// TIA Portal project "HydroPlantProject_V15.1" (V15.1) (continued)

   IF "StationIntHoa" = 1 OR ("StationIntHoa" = 2 AND "StationIntl_Ctrl") THEN
       "StationInterlock_Out" := 1;
   END_IF;

   IF "BaffleHOA" = 0 OR ("BaffleHOA" = 2 AND NOT "Baffle_Ctrl") THEN
       "Baffle_En" := 0;
   END_IF;

   IF "BaffleHOA" = 1 OR ("BaffleHOA" = 2 AND "Baffle_Ctrl") THEN
       "Baffle_En" := 1;
   END_IF;





   //Analog Outputs
   "SCP"(Input_Min:=0,
         Input_Signal:="OilPumpVFDpct",
         Input_Max:=100,
         Output_Min:=0,
         Output_Max:=27648,
         SV=>"OilPumpVFDsp_Out");

   "SCP"(Input_Min := 0,
         Input_Signal := "BafflePct",
         Input_Max := 100,
         Output_Min := 0,
         Output_Max := 27648,
         SV => "Baffle_Out");


   //Analog Inputs
   "SCP"(Input_Min:=0,
         Input_Signal:="OilTemp_In",
         Input_Max:=27648,
         Output_Min:=0,
         Output_Max:=500,
         SV=>"OilTemp");

   "SCP"(Input_Min := 0,
         Input_Signal := "OilFlow_In",
         Input_Max := 27648,
         Output_Min := 0,
         Output_Max := 30,
         SV => "OilFlow");

   "SCP"(Input_Min := 0,
         Input_Signal := "RPM_In",
   Input_Max := 27648,
   Output_Min := 0,
   Output_Max := 200,
   SV => "RPM");

   "SCP"(Input_Min := 0,
         Input_Signal := "Current_In",
         Input_Max := 27648,
         Output_Min := 0,
         Output_Max := 700,
         SV => "Current");


   //Full Auto Bit
   IF "BaffleHOA" = 2 AND "AlarmHornHoa" = 0 AND "VFDHOA" = 0 AND "StationIntHoa" = 0 AND "BrakeHoa" = 0 THEN
       "FullAutoBit" := 1;
   ELSE
       "FullAutoBit" := 0;
   END_IF;
END_FUNCTION_BLOCK

FUNCTION_BLOCK "IO_STL"   // FB5, STL
{ S7_Optimized_Access := 'TRUE' }
VERSION : 0.1
BEGIN

REGION Network 1
   //Digital Outputs
         A     "OilLowFlowAlarm";
         JC    ResetOilPumpVFD;
         CLR;
         A     "EStopAlarm";
         JC    ResetOilPumpVFD;
         L     "VFDHOA";
         L     0;
         ==I;
         JC    ResetOilPumpVFD;
         CLR;
         L     "VFDHOA";
         L     1;
         ==I;
         JC    SetOilPumpVFD;
         CLR;
         L     "VFDHOA";
         L     2;
         ==I;
         JC    AutoOilPumpVFD;

   AutoOilPumpVFD:A     "OilPumpVFD_Ctrl";
         JC    SetOilPumpVFD;
         JU    ResetOilPumpVFD;

   SetOilPumpVFD:AN    "OilLowFlowAlarm";
         AN    "EStop";
         S     "OilPumpVFDen_Out";
         JU    Brake;

   ResetOilPumpVFD:R     "OilPumpVFDen_Out";
         JU    Brake;

   Brake:L     "BrakeHoa";
         L     0;
         ==I;
         JC    ResetBrake;
         CLR;
         L     "BrakeHoa";
         L     1;
         ==I;
         JC    SetBrake;
         CLR;
         L     "BrakeHoa";
         L     2;
         ==I;
         JC    AutoBrake;

   AutoBrake:A     "Brake_Ctrl";
         JC    SetBrake;
         JU    ResetBrake;

   SetBrake:S     "Brake_Out";
         JU    AlarmHorn;

   ResetBrake:R     "Brake_Out";
         JU    AlarmHorn;

   AlarmHorn:L     "AlarmHornHoa";
         L     0;
         ==I;
         JC    ResetAlarmHorn;
         CLR;
         L     "AlarmHornHoa";
         L     1;
         ==I;
         JC    SetAlarmHorn;
         CLR;
         L     "AlarmHornHoa";
         L     2;
         ==I;
         JC    AutoAlarmHorn;

   AutoAlarmHorn:A     "AlarmHorn_Ctrl";
         JC    SetAlarmHorn;
         JU    ResetAlarmHorn;

   SetAlarmHorn:S     "AlarmHorn_Out";
         JU    StationInterlock;

   ResetAlarmHorn:R     "AlarmHorn_Out";
         JU    StationInterlock;

   StationInterlock:A     "EStopAlarm";
         JC    ResetStationInterlock;
         L     "StationIntHoa";
         L     0;
         ==I;
         JC    ResetStationInterlock;
         CLR;
         L     "StationIntHoa";
         L     1;
         ==I;
         JC    SetStationInterlock;
         CLR;
         L     "StationIntHoa";
         L     2;
         ==I;
         JC    AutoStationInterlock;

   AutoStationInterlock:A     "StationIntl_Ctrl";
         JC    SetStationInterlock;
         JU    ResetStationInterlock;

   SetStationInterlock:AN    "EStopAlarm";
         S     "StationInterlock_Out";
         JU    Baffle;

   ResetStationInterlock:R     "StationInterlock_Out";
         JU    Baffle;

   Baffle:L     "BaffleHOA";
         L     0;
         ==I;
         JC    ResetBaffle;
         CLR;
         L     "BaffleHOA";
         L     1;
         ==I;
         JC    SetBaffle;
         CLR;
         L     "BaffleHOA";
         L     2;
         ==I;
         JC    AutoBaffle;

   AutoBaffle:A     "Baffle_Ctrl";
         JC    SetBaffle;
         JU    ResetBaffle;

   SetBaffle:S     "Baffle_En";
         JU    AnalogOutputs;

   ResetBaffle:R     "Baffle_En";
         JU    AnalogOutputs;



   //Analog Outputs
   AnalogOutputs:CALL  "SCP"
         ( Input_Min    := 0,
           Input_Signal := "OilPumpVFDpct",
           Input_Max    := 100,
           Output_Min   := 0,
           Output_Max   := 27648,
           SV           := "OilPumpVFDsp_Out"
         );
         JU    AnalogInputs;

         CALL  "SCP"
         ( Input_Min    := 0,
           Input_Signal := "BafflePct",
           Input_Max    := 100,
           Output_Min   := 0,
           Output_Max   := 27648,
           SV           := "Baffle_Out"
         );


   //Analog Inputs
   AnalogInputs:CALL  "SCP"
         ( Input_Min    := 0,
           Input_Signal := "OilTemp_In",
           Input_Max    := 27648,
           Output_Min   := 0,
           Output_Max   := 500,
           SV           := "OilTemp"
         );

         CALL  "SCP"
         ( Input_Min    := 0,
           Input_Signal := "OilFlow_In",
           Input_Max    := 27648,
           Output_Min   := 0,
           Output_Max   := 30,
           SV           := "OilFlow"
         );

         CALL  "SCP"
         ( Input_Min    := 0,
           Input_Signal := "RPM_In",
           Input_Max    := 27648,
           Output_Min   := 0,
           Output_Max   := 200,
           SV           := "RPM"
         );

         CALL  "SCP"
         ( Input_Min    := 0,
           Input_Signal := "Current_In",
           Input_Max    := 27648,
           Output_Min   := 0,
           Output_Max   := 700,
           SV           := "Current"
         );

   //Full Auto Bit
         CLR;
         L     "BaffleHOA";
         L     2;
         ==I;
         NOT;
         JC    ResetFullAuto;
         CLR;
         L     "VFDHOA";
         L     2;
         ==I;
         NOT;
         JC    ResetFullAuto;
         CLR;
         L     "AlarmHornHoa";
         L     2;
         ==I;
         NOT;
         JC    ResetFullAuto;
         CLR;
         L     "BrakeHoa";
         L     2;
         ==I;
         NOT;
         JC    ResetFullAuto;
         CLR;
         L     "StationIntHoa";
         L     2;
         ==I;
         NOT;
         JC    ResetFullAuto;
         CLR;
         SET;
         S     "FullAutoBit";
         JU    EndOfLine;

   ResetFullAuto:SET;
         NOT;
         R     "FullAutoBit";
         JU    EndOfLine;

   EndOfLine:BE;
END_REGION
END_FUNCTION_BLOCK

FUNCTION_BLOCK "ALARMS_LAD"   // FB6, LAD
{ S7_Optimized_Access := 'TRUE' }
VERSION : 0.1
   VAR
      OS1 : Bool;
      OS2 : Bool;
      OS3 : Bool;
      OS4 : Bool;
      OS5 : Bool;
      OS6 : Bool;
      OS7 : Bool;
      OS8 : Bool;
   END_VAR
   VAR_TEMP
      tv : Time;
      Tsp : Int;
      OLFAT : Bool;
      OLFD : Int;
      tv1 : Time;
      OCD : Int;
      tv2 : Time;
      OCAT : Bool;
      HOTD : Int;
      tv3 : Time;
      HOTAT : Bool;
      OSD : Int;
      tv4 : Time;
      OSAT : Bool;
      OHFD : Int;
      tv5 : Time;
      OHFAT : Bool;
      BFD : Int;
      tv6 : Time;
      BFAT : Bool;
      ESAT : Bool;
      AlarmHornTrigger : Bool;
   END_VAR
   VAR_TEMP   // added for the SCL form of the ladder/FBD networks
      _w1 : Bool;
      _w2 : Bool;
   END_VAR
BEGIN

REGION Network 1
   // Oil Low Flow Alarm
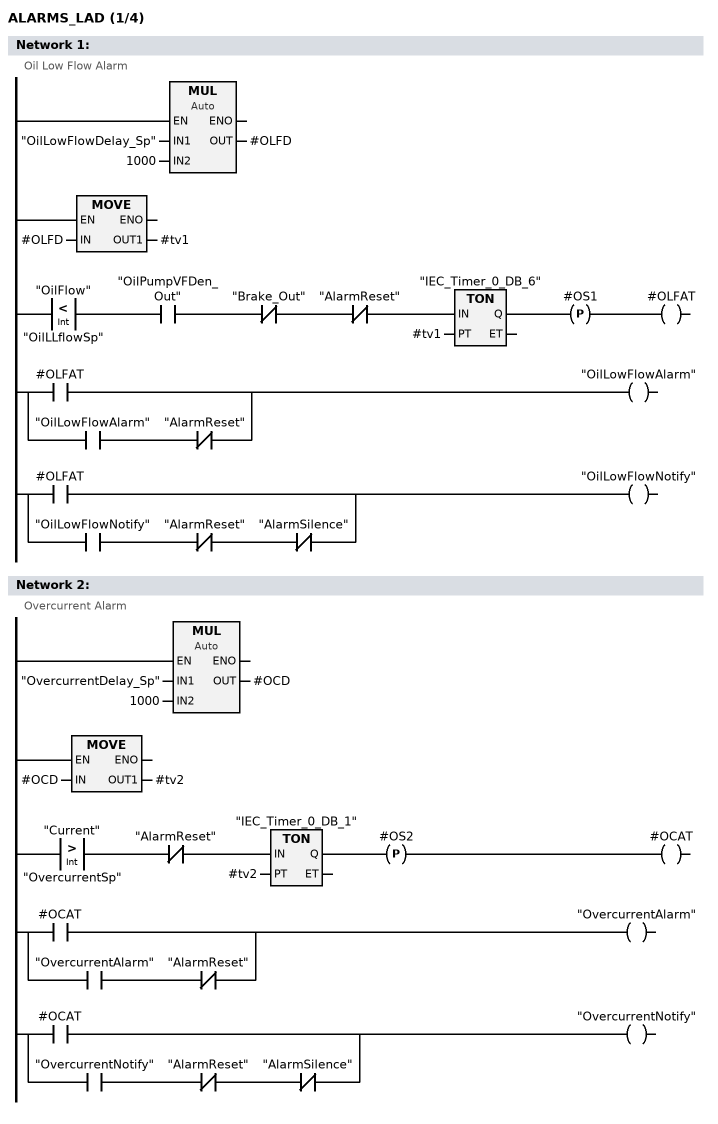
   #OLFD := "OilLowFlowDelay_Sp" * 1000;
   #tv1 := #OLFD;
   "IEC_Timer_0_DB_6".TON(IN := ("OilFlow" < "OilLLflowSp") AND "OilPumpVFDen_Out" AND NOT "Brake_Out" AND NOT "AlarmReset",
                          PT := #tv1);
   #_w1 := "IEC_Timer_0_DB_6".Q AND NOT #OS1;   // rising edge
   #OS1 := "IEC_Timer_0_DB_6".Q;
   #OLFAT := #_w1;
   "OilLowFlowAlarm" := #OLFAT OR ("OilLowFlowAlarm" AND NOT "AlarmReset");
   "OilLowFlowNotify" := #OLFAT OR ("OilLowFlowNotify" AND NOT "AlarmReset" AND NOT "AlarmSilence");
END_REGION

REGION Network 2
   // Overcurrent Alarm
   #OCD := "OvercurrentDelay_Sp" * 1000;
   #tv2 := #OCD;
   "IEC_Timer_0_DB_1".TON(IN := ("Current" > "OvercurrentSp") AND NOT "AlarmReset", PT := #tv2);
   #_w1 := "IEC_Timer_0_DB_1".Q AND NOT #OS2;   // rising edge
   #OS2 := "IEC_Timer_0_DB_1".Q;
   #OCAT := #_w1;
   "OvercurrentAlarm" := #OCAT OR ("OvercurrentAlarm" AND NOT "AlarmReset");
   "OvercurrentNotify" := #OCAT OR ("OvercurrentNotify" AND NOT "AlarmReset" AND NOT "AlarmSilence");
END_REGION

REGION Network 3
   // High Oil Temp Alarm
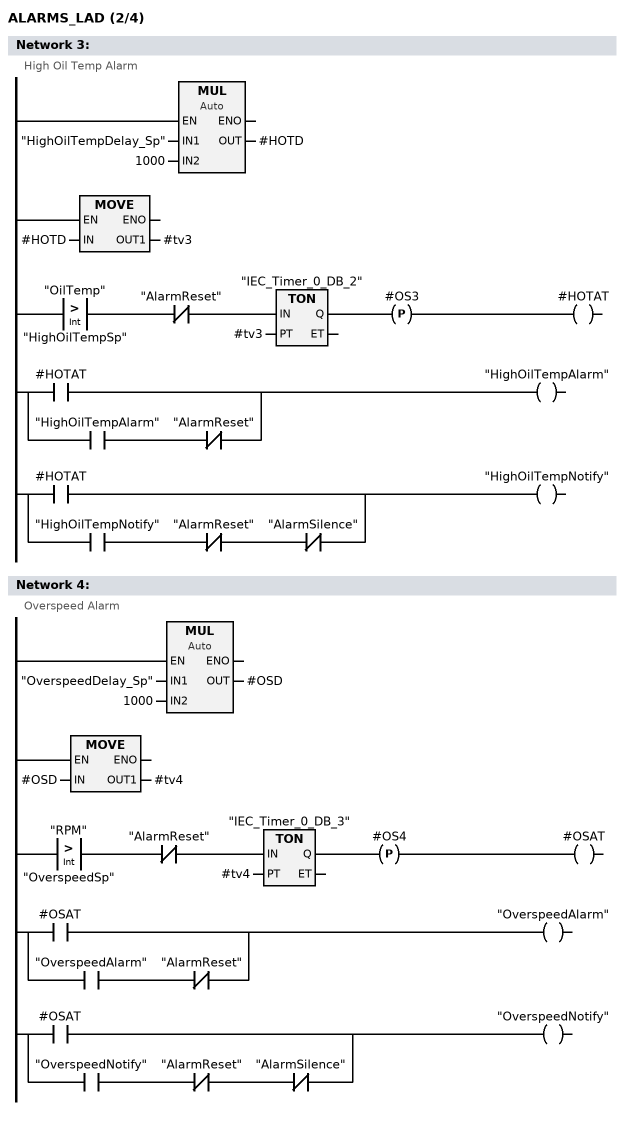
   #HOTD := "HighOilTempDelay_Sp" * 1000;
   #tv3 := #HOTD;
   "IEC_Timer_0_DB_2".TON(IN := ("OilTemp" > "HighOilTempSp") AND NOT "AlarmReset", PT := #tv3);
   #_w1 := "IEC_Timer_0_DB_2".Q AND NOT #OS3;   // rising edge
   #OS3 := "IEC_Timer_0_DB_2".Q;
   #HOTAT := #_w1;
   "HighOilTempAlarm" := #HOTAT OR ("HighOilTempAlarm" AND NOT "AlarmReset");
   "HighOilTempNotify" := #HOTAT OR ("HighOilTempNotify" AND NOT "AlarmReset" AND NOT "AlarmSilence");
END_REGION

REGION Network 4
   // Overspeed Alarm
   #OSD := "OverspeedDelay_Sp" * 1000;
   #tv4 := #OSD;
   "IEC_Timer_0_DB_3".TON(IN := ("RPM" > "OverspeedSp") AND NOT "AlarmReset", PT := #tv4);
   #_w1 := "IEC_Timer_0_DB_3".Q AND NOT #OS4;   // rising edge
   #OS4 := "IEC_Timer_0_DB_3".Q;
   #OSAT := #_w1;
   "OverspeedAlarm" := #OSAT OR ("OverspeedAlarm" AND NOT "AlarmReset");
   "OverspeedNotify" := #OSAT OR ("OverspeedNotify" AND NOT "AlarmReset" AND NOT "AlarmSilence");
END_REGION

REGION Network 5
   // Oil High Flow Alarm
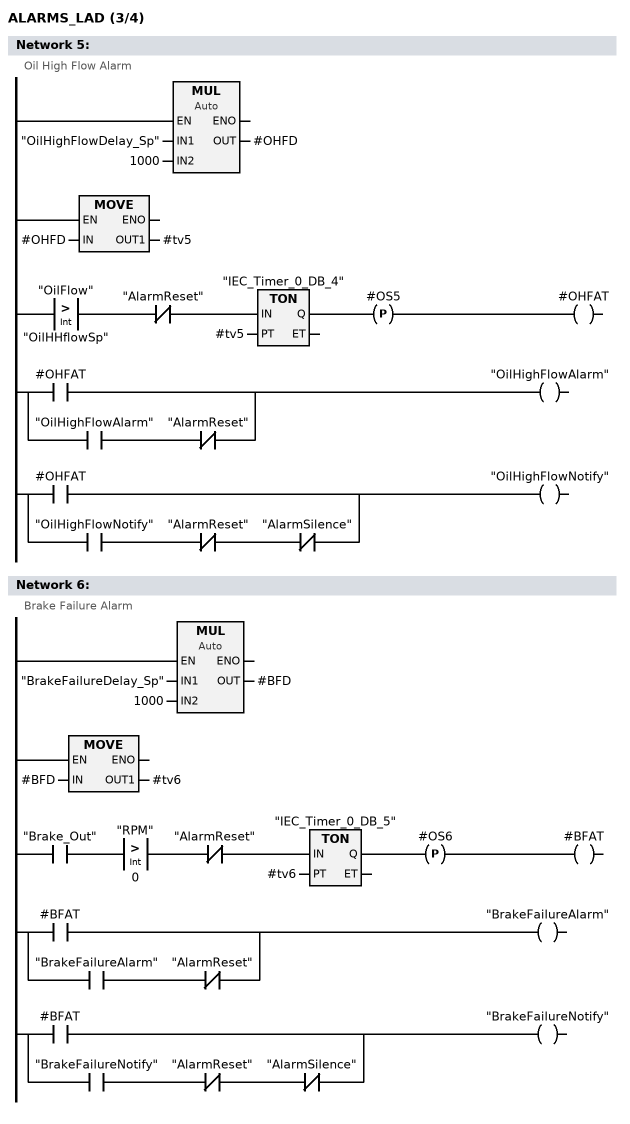
   #OHFD := "OilHighFlowDelay_Sp" * 1000;
   #tv5 := #OHFD;
   "IEC_Timer_0_DB_4".TON(IN := ("OilFlow" > "OilHHflowSp") AND NOT "AlarmReset", PT := #tv5);
   #_w1 := "IEC_Timer_0_DB_4".Q AND NOT #OS5;   // rising edge
   #OS5 := "IEC_Timer_0_DB_4".Q;
   #OHFAT := #_w1;
   "OilHighFlowAlarm" := #OHFAT OR ("OilHighFlowAlarm" AND NOT "AlarmReset");
   "OilHighFlowNotify" := #OHFAT OR ("OilHighFlowNotify" AND NOT "AlarmReset" AND NOT "AlarmSilence");
END_REGION

REGION Network 6
   // Brake Failure Alarm
   #BFD := "BrakeFailureDelay_Sp" * 1000;
   #tv6 := #BFD;
   "IEC_Timer_0_DB_5".TON(IN := "Brake_Out" AND ("RPM" > 0) AND NOT "AlarmReset", PT := #tv6);
   #_w1 := "IEC_Timer_0_DB_5".Q AND NOT #OS6;   // rising edge
   #OS6 := "IEC_Timer_0_DB_5".Q;
   #BFAT := #_w1;
   "BrakeFailureAlarm" := #BFAT OR ("BrakeFailureAlarm" AND NOT "AlarmReset");
   "BrakeFailureNotify" := #BFAT OR ("BrakeFailureNotify" AND NOT "AlarmReset" AND NOT "AlarmSilence");
END_REGION

REGION Network 7
   // EStop Alarm
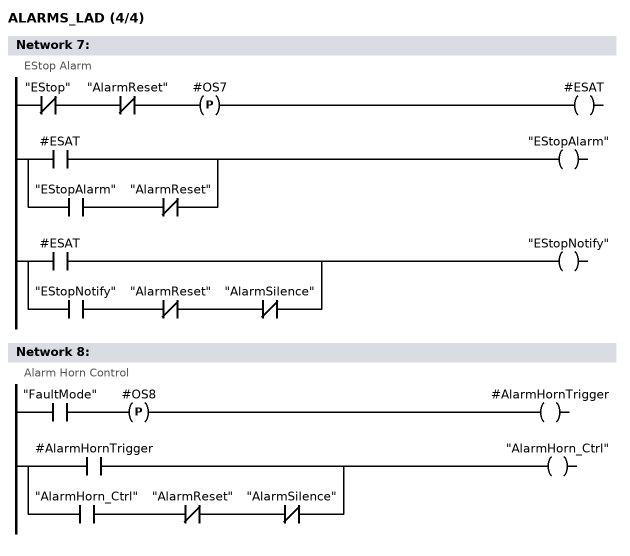
   RUNG wire#powerrail
      I_Contact( "EStop" )
      I_Contact( "AlarmReset" )
      P_Trig( #OS7 )
      Coil( #ESAT )
   END_RUNG
   RUNG wire#powerrail
      Contact( #ESAT )
      wire#w1
      Coil( "EStopAlarm" )
   END_RUNG
   RUNG wire#powerrail
      Contact( "EStopAlarm" )
      I_Contact( "AlarmReset" )
   END_RUNG wire#w1
   RUNG wire#powerrail
      Contact( #ESAT )
      wire#w2
      Coil( "EStopNotify" )
   END_RUNG
   RUNG wire#powerrail
      Contact( "EStopNotify" )
      I_Contact( "AlarmReset" )
      I_Contact( "AlarmSilence" )
   END_RUNG wire#w2
   // the same network as SCL:
   #_w1 := NOT "EStop" AND NOT "AlarmReset";
   #_w2 := #_w1 AND NOT #OS7;   // rising edge
   #OS7 := #_w1;
   #ESAT := #_w2;
   "EStopAlarm" := #ESAT OR ("EStopAlarm" AND NOT "AlarmReset");
   "EStopNotify" := #ESAT OR ("EStopNotify" AND NOT "AlarmReset" AND NOT "AlarmSilence");
END_REGION

REGION Network 8
   // Alarm Horn Control
   RUNG wire#powerrail
      Contact( "FaultMode" )
      P_Trig( #OS8 )
      Coil( #AlarmHornTrigger )
   END_RUNG
   RUNG wire#powerrail
      Contact( #AlarmHornTrigger )
      wire#w1
      Coil( "AlarmHorn_Ctrl" )
   END_RUNG
   RUNG wire#powerrail
      Contact( "AlarmHorn_Ctrl" )
      I_Contact( "AlarmReset" )
      I_Contact( "AlarmSilence" )
   END_RUNG wire#w1
   // the same network as SCL:
   #_w1 := "FaultMode" AND NOT #OS8;   // rising edge
   #OS8 := "FaultMode";
   #AlarmHornTrigger := #_w1;
   "AlarmHorn_Ctrl" := #AlarmHornTrigger OR ("AlarmHorn_Ctrl" AND NOT "AlarmReset" AND NOT "AlarmSilence");
END_REGION
END_FUNCTION_BLOCK

FUNCTION_BLOCK "HOA_FBD"   // FB7, FBD
{ S7_Optimized_Access := 'TRUE' }
VERSION : 0.1
   VAR
      OS1 : Bool;
      OS3 : Bool;
      OS2 : Bool;
      OS4 : Bool;
      OS5 : Bool;
      OS6 : Bool;
      OS7 : Bool;
      OS8 : Bool;
      OS9 : Bool;
      OS10 : Bool;
      OS11 : Bool;
      OS12 : Bool;
   END_VAR
   VAR_TEMP   // added for the SCL form of the ladder/FBD networks
      _w1 : Bool;
      _w2 : Bool;
      _w3 : Bool;
   END_VAR
BEGIN

REGION Network 1
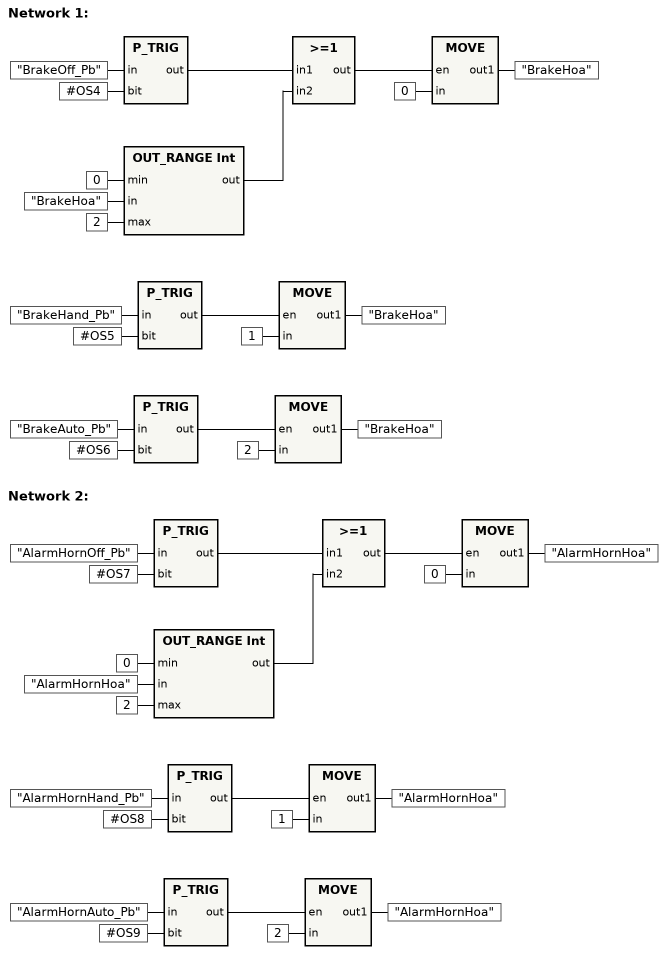
   #_w1 := "BrakeOff_Pb" AND NOT #OS4;   // rising edge
   #OS4 := "BrakeOff_Pb";
   IF #_w1 OR ("BrakeHoa" < 0) OR ("BrakeHoa" > 2) THEN "BrakeHoa" := 0; END_IF;
   #_w2 := "BrakeHand_Pb" AND NOT #OS5;   // rising edge
   #OS5 := "BrakeHand_Pb";
   IF #_w2 THEN "BrakeHoa" := 1; END_IF;
   #_w3 := "BrakeAuto_Pb" AND NOT #OS6;   // rising edge
   #OS6 := "BrakeAuto_Pb";
   IF #_w3 THEN "BrakeHoa" := 2; END_IF;
END_REGION

REGION Network 2
   #_w1 := "AlarmHornOff_Pb" AND NOT #OS7;   // rising edge
   #OS7 := "AlarmHornOff_Pb";
   IF #_w1 OR ("AlarmHornHoa" < 0) OR ("AlarmHornHoa" > 2) THEN "AlarmHornHoa" := 0; END_IF;
   #_w2 := "AlarmHornHand_Pb" AND NOT #OS8;   // rising edge
   #OS8 := "AlarmHornHand_Pb";
   IF #_w2 THEN "AlarmHornHoa" := 1; END_IF;
   #_w3 := "AlarmHornAuto_Pb" AND NOT #OS9;   // rising edge
   #OS9 := "AlarmHornAuto_Pb";
   IF #_w3 THEN "AlarmHornHoa" := 2; END_IF;
END_REGION

REGION Network 3
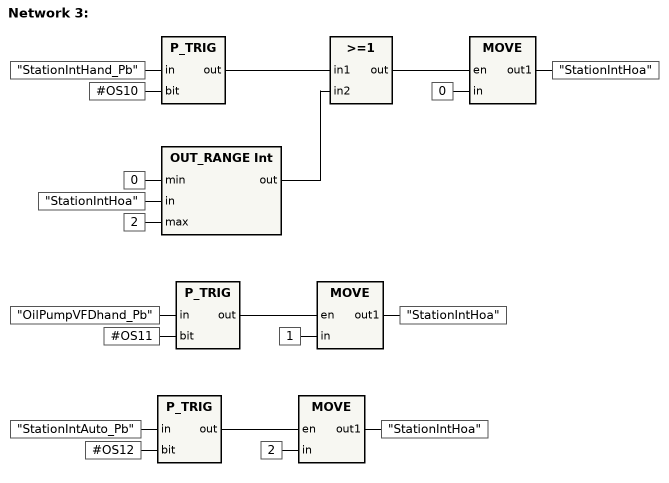
   #_w1 := "StationIntHand_Pb" AND NOT #OS10;   // rising edge
   #OS10 := "StationIntHand_Pb";
   IF #_w1 OR ("StationIntHoa" < 0) OR ("StationIntHoa" > 2) THEN "StationIntHoa" := 0; END_IF;
   #_w2 := "OilPumpVFDhand_Pb" AND NOT #OS11;   // rising edge
   #OS11 := "OilPumpVFDhand_Pb";
   IF #_w2 THEN "StationIntHoa" := 1; END_IF;
   #_w3 := "StationIntAuto_Pb" AND NOT #OS12;   // rising edge
   #OS12 := "StationIntAuto_Pb";
   IF #_w3 THEN "StationIntHoa" := 2; END_IF;
END_REGION
END_FUNCTION_BLOCK

FUNCTION_BLOCK "HOA_LAD"   // FB8, LAD
{ S7_Optimized_Access := 'TRUE' }
VERSION : 0.1
   VAR
      OS1 : Bool;
      OS2 : Bool;
      OS3 : Bool;
      OS4 : Bool;
      OS5 : Bool;
      OS6 : Bool;
      OS7 : Bool;
      OS8 : Bool;
      OS9 : Bool;
      OS10 : Bool;
      OS11 : Bool;
      OS12 : Bool;
   END_VAR
   VAR_TEMP   // added for the SCL form of the ladder/FBD networks
      _w1 : Bool;
      _w2 : Bool;
      _w3 : Bool;
   END_VAR
BEGIN

REGION Network 1
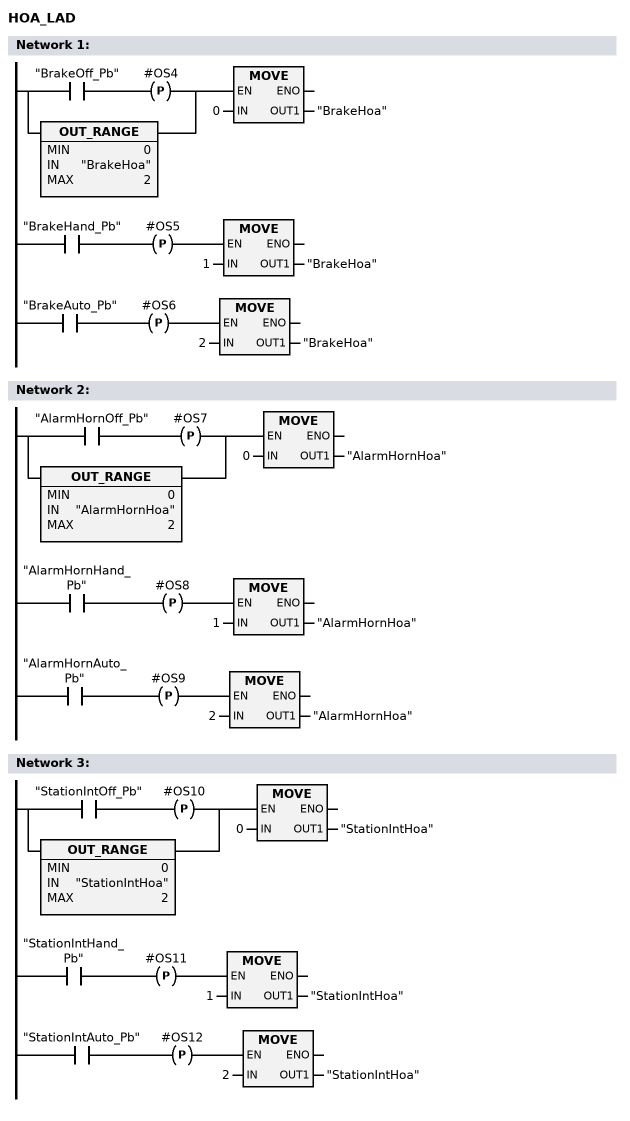
   #_w1 := "BrakeOff_Pb" AND NOT #OS4;   // rising edge
   #OS4 := "BrakeOff_Pb";
   IF #_w1 OR ("BrakeHoa" < 0) OR ("BrakeHoa" > 2) THEN "BrakeHoa" := 0; END_IF;
   #_w2 := "BrakeHand_Pb" AND NOT #OS5;   // rising edge
   #OS5 := "BrakeHand_Pb";
   IF #_w2 THEN "BrakeHoa" := 1; END_IF;
   #_w3 := "BrakeAuto_Pb" AND NOT #OS6;   // rising edge
   #OS6 := "BrakeAuto_Pb";
   IF #_w3 THEN "BrakeHoa" := 2; END_IF;
END_REGION

REGION Network 2
   #_w1 := "AlarmHornOff_Pb" AND NOT #OS7;   // rising edge
   #OS7 := "AlarmHornOff_Pb";
   IF #_w1 OR ("AlarmHornHoa" < 0) OR ("AlarmHornHoa" > 2) THEN "AlarmHornHoa" := 0; END_IF;
   #_w2 := "AlarmHornHand_Pb" AND NOT #OS8;   // rising edge
   #OS8 := "AlarmHornHand_Pb";
   IF #_w2 THEN "AlarmHornHoa" := 1; END_IF;
   #_w3 := "AlarmHornAuto_Pb" AND NOT #OS9;   // rising edge
   #OS9 := "AlarmHornAuto_Pb";
   IF #_w3 THEN "AlarmHornHoa" := 2; END_IF;
END_REGION

REGION Network 3
   #_w1 := "StationIntOff_Pb" AND NOT #OS10;   // rising edge
   #OS10 := "StationIntOff_Pb";
   IF #_w1 OR ("StationIntHoa" < 0) OR ("StationIntHoa" > 2) THEN "StationIntHoa" := 0; END_IF;
   #_w2 := "StationIntHand_Pb" AND NOT #OS11;   // rising edge
   #OS11 := "StationIntHand_Pb";
   IF #_w2 THEN "StationIntHoa" := 1; END_IF;
   #_w3 := "StationIntAuto_Pb" AND NOT #OS12;   // rising edge
   #OS12 := "StationIntAuto_Pb";
   IF #_w3 THEN "StationIntHoa" := 2; END_IF;
END_REGION
END_FUNCTION_BLOCK

FUNCTION_BLOCK "HOA_SCL"   // FB9, SCL
{ S7_Optimized_Access := 'TRUE' }
VERSION : 0.1
BEGIN
   //Brake HOA Controls
   IF "BrakeHoa" < 0 OR "BrakeHoa" > 2 THEN
       "BrakeHoa" := 0;
   END_IF;

   IF "BrakeOff_Pb" AND "BrakeHoa" <> 0 THEN
       "BrakeHoa" := 0;
   END_IF;

   IF "BrakeHand_Pb" AND "BrakeHoa" <> 1 THEN
       "BrakeHoa" := 1;
   END_IF;

   IF "BrakeAuto_Pb" AND "BrakeHoa" <> 2 THEN
       "BrakeHoa" := 2;
   END_IF;


   //Alarm Horn HOA Controls
   IF "AlarmHornHoa" < 0 OR "AlarmHornHoa" > 2 THEN
       "AlarmHornHoa" := 0;
   END_IF;

   IF "AlarmHornOff_Pb" AND "AlarmHornHoa" <> 0 THEN
       "AlarmHornHoa" := 0;
   END_IF;

   IF "AlarmHornHand_Pb" AND "AlarmHornHoa" <> 1 THEN
       "AlarmHornHoa" := 1;
   END_IF;

   IF "AlarmHornAuto_Pb" AND "AlarmHornHoa" <> 2 THEN
       "AlarmHornHoa" := 2;
   END_IF;


   //Station Interlock HOA Controls
   IF "StationIntHoa" < 0 OR "StationIntHoa" > 2 THEN
       "StationIntHoa" := 0;
   END_IF;

   IF "StationIntOff_Pb" AND "StationIntHoa" <> 0 THEN
       "StationIntHoa" := 0;
   END_IF;

   IF "StationIntHand_Pb" AND "StationIntHoa" <> 1 THEN
       "StationIntHoa" := 1;
   END_IF;

   IF "StationIntAuto_Pb" AND "StationIntHoa" <> 2 THEN
       "StationIntHoa" := 2;
   END_IF;
END_FUNCTION_BLOCK

FUNCTION_BLOCK "HOA_STL"   // FB10, STL
{ S7_Optimized_Access := 'TRUE' }
VERSION : 0.1
   VAR
      OS1 : Bool;
      OS2 : Bool;
      OS4 : Bool;
      OS5 : Bool;
      OS12 : Bool;
      OS6 : Bool;
      OS7 : Bool;
      OS8 : Bool;
      OS9 : Bool;
      OS10 : Bool;
      OS11 : Bool;
      OS3 : Bool;
   END_VAR
BEGIN

REGION Network 1
         L     "BrakeHoa";
         L     0;
         <I;
         JC    SetBrakeHoaZero;
         CLR;
         L     "BrakeHoa";
         L     2;
         >I;
         JC    SetBrakeHoaZero;
         CLR;
         A     "BrakeOff_Pb";
         FP    #OS4;
         JC    SetBrakeHoaZero;
         CLR;
         A     "BrakeHand_Pb";
         FP    #OS5;
         JC    SetBrakeHoaOne;
         CLR;
         A     "BrakeAuto_Pb";
         FP    #OS6;
         JC    SetBrakeHoaTwo;
         JU    AlarmHorn;

   SetBrakeHoaZero:L     0;
         T     "BrakeHoa";
         JU    AlarmHorn;

   SetBrakeHoaOne:L     1;
         T     "BrakeHoa";
         JU    AlarmHorn;

   SetBrakeHoaTwo:L     2;
         T     "BrakeHoa";
         JU    AlarmHorn;


   AlarmHorn:L     "AlarmHornHoa";
         L     0;
         <I;
         JC    SetAlarmHornHoaZero;
         CLR;
         L     "AlarmHornHoa";
         L     2;
         >I;
         JC    SetAlarmHornHoaZero;
         CLR;
         A     "AlarmHornOff_Pb";
         FP    #OS7;
         JC    SetAlarmHornHoaZero;
         CLR;
         A     "AlarmHornHand_Pb";
         FP    #OS8;
         JC    SetBrakeHoaOne;
         CLR;
         A     "AlarmHornAuto_Pb";
         FP    #OS9;
         JC    SetOAlarmHornHoaTwo;
         JU    StationInterlock;

   SetAlarmHornHoaZero:L     0;
         T     "AlarmHornHoa";
         JU    StationInterlock;

   SetOAlarmHornHoaOne:L     1;
         T     "AlarmHornHoa";
         JU    StationInterlock;

   SetOAlarmHornHoaTwo:L     2;
         T     "AlarmHornHoa";
         JU    StationInterlock;


   StationInterlock:L     "StationIntHoa";
         L     0;
         <I;
         JC    SetStationInterlockHoaZero;
         CLR;
         L     "StationIntHoa";
         L     2;
         >I;
         JC    SetStationInterlockHoaZero;
         CLR;
         A     "StationIntOff_Pb";
         FP    #OS10;
         JC    SetStationInterlockHoaZero;
         CLR;
         A     "StationIntHand_Pb";
         FP    #OS11;
         JC    SetStationInterlockHoaOne;
         CLR;
         A     "StationIntAuto_Pb";
         FP    #OS12;
         JC    SetStationInterlockHoaTwo;
         JU    EndOfLine;

   SetStationInterlockHoaZero:L     0;
         T     "StationIntHoa";
         BE;

   SetStationInterlockHoaOne:L     1;
         T     "StationIntHoa";
         BE;

   SetStationInterlockHoaTwo:L     2;
         T     "StationIntHoa";
         BE;

   EndOfLine:BE;
END_REGION
END_FUNCTION_BLOCK

FUNCTION_BLOCK "ALARMS_FBD"   // FB11, FBD
{ S7_Optimized_Access := 'TRUE' }
VERSION : 0.1
   VAR
      OS1 : Bool;
      OS2 : Bool;
      OS3 : Bool;
      OS4 : Bool;
      OS5 : Bool;
      OS6 : Bool;
      OS7 : Bool;
   END_VAR
   VAR_TEMP
      ti1 : Int;
      tt1 : Time;
      ti2 : Int;
      tt2 : Time;
      ti3 : Int;
      tt3 : Time;
      ti4 : Int;
      tt4 : Time;
      ti5 : Int;
      tt5 : Time;
      ti6 : Int;
      tt6 : Time;
   END_VAR
   VAR_TEMP   // added for the SCL form of the ladder/FBD networks
      _w1 : Bool;
   END_VAR
BEGIN

REGION Network 1
   // Oil Low Flow Alarm
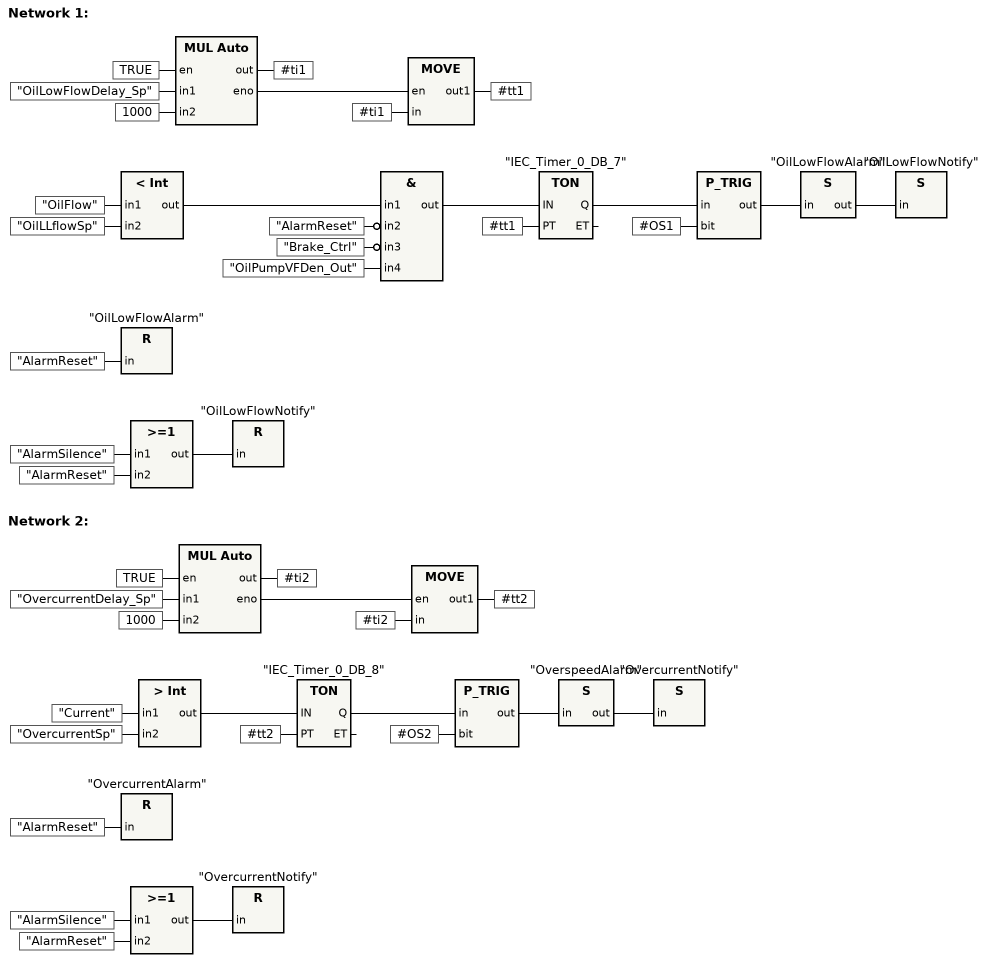
   IF TRUE THEN
       #ti1 := "OilLowFlowDelay_Sp" * 1000;
       #tt1 := #ti1;
   END_IF;
   "IEC_Timer_0_DB_7".TON(IN := ("OilFlow" < "OilLLflowSp") AND NOT "AlarmReset" AND NOT "Brake_Ctrl" AND "OilPumpVFDen_Out",
                          PT := #tt1);
   #_w1 := "IEC_Timer_0_DB_7".Q AND NOT #OS1;   // rising edge
   #OS1 := "IEC_Timer_0_DB_7".Q;
   IF #_w1 THEN
       "OilLowFlowAlarm" := TRUE;
       "OilLowFlowNotify" := TRUE;
   END_IF;
   IF "AlarmReset" THEN "OilLowFlowAlarm" := FALSE; END_IF;
   IF "AlarmSilence" OR "AlarmReset" THEN "OilLowFlowNotify" := FALSE; END_IF;
END_REGION

REGION Network 2
   // Overcurrent Alarm
   IF TRUE THEN
       #ti2 := "OvercurrentDelay_Sp" * 1000;
       #tt2 := #ti2;
   END_IF;
   "IEC_Timer_0_DB_8".TON(IN := "Current" > "OvercurrentSp", PT := #tt2);
   #_w1 := "IEC_Timer_0_DB_8".Q AND NOT #OS2;   // rising edge
   #OS2 := "IEC_Timer_0_DB_8".Q;
   IF #_w1 THEN
       "OverspeedAlarm" := TRUE;
       "OvercurrentNotify" := TRUE;
   END_IF;
   IF "AlarmReset" THEN "OvercurrentAlarm" := FALSE; END_IF;
   IF "AlarmSilence" OR "AlarmReset" THEN "OvercurrentNotify" := FALSE; END_IF;
END_REGION

REGION Network 3
   // High Oil Temp Alarm
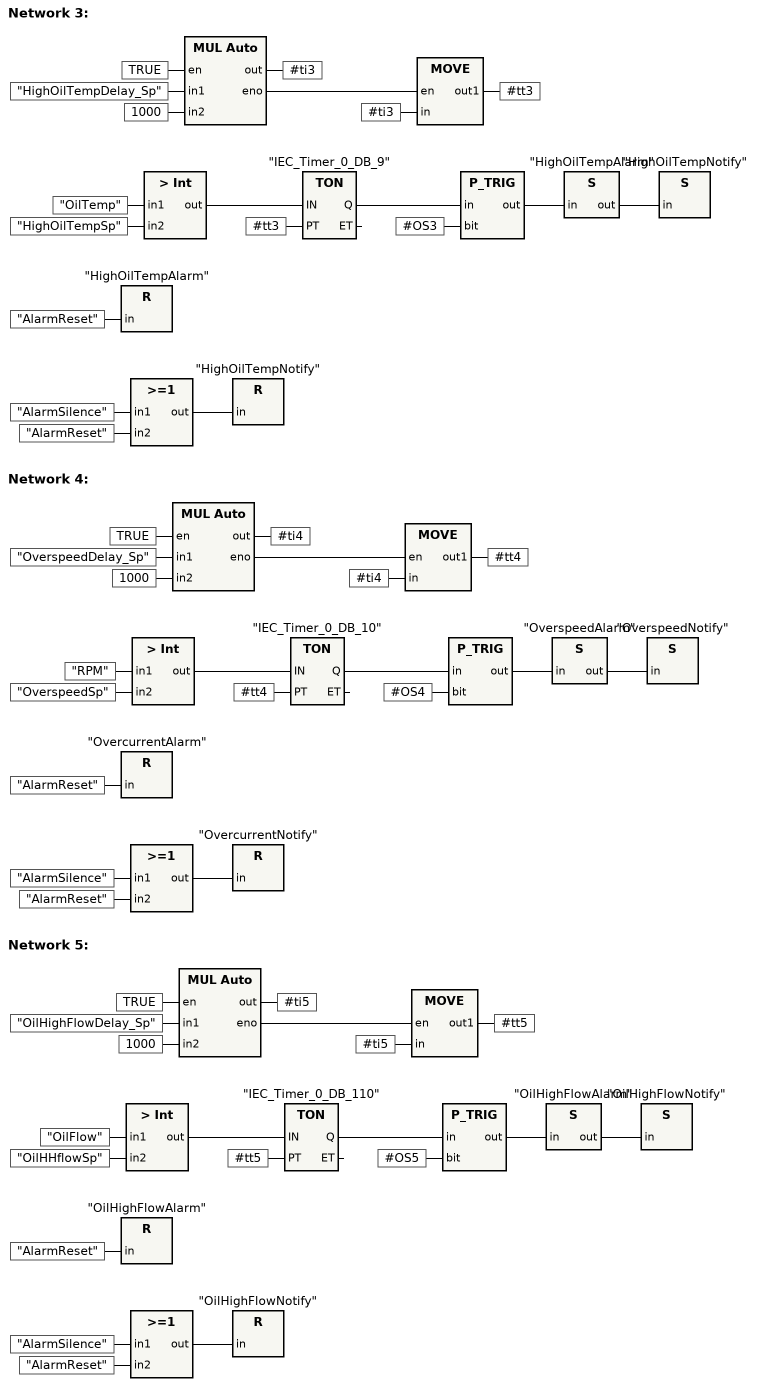
   IF TRUE THEN
       #ti3 := "HighOilTempDelay_Sp" * 1000;
       #tt3 := #ti3;
   END_IF;
   "IEC_Timer_0_DB_9".TON(IN := "OilTemp" > "HighOilTempSp", PT := #tt3);
   #_w1 := "IEC_Timer_0_DB_9".Q AND NOT #OS3;   // rising edge
   #OS3 := "IEC_Timer_0_DB_9".Q;
   IF #_w1 THEN
       "HighOilTempAlarm" := TRUE;
       "HighOilTempNotify" := TRUE;
   END_IF;
   IF "AlarmReset" THEN "HighOilTempAlarm" := FALSE; END_IF;
   IF "AlarmSilence" OR "AlarmReset" THEN "HighOilTempNotify" := FALSE; END_IF;
END_REGION

REGION Network 4
   // Overspeed Alarm
   IF TRUE THEN
       #ti4 := "OverspeedDelay_Sp" * 1000;
       #tt4 := #ti4;
   END_IF;
   "IEC_Timer_0_DB_10".TON(IN := "RPM" > "OverspeedSp", PT := #tt4);
   #_w1 := "IEC_Timer_0_DB_10".Q AND NOT #OS4;   // rising edge
   #OS4 := "IEC_Timer_0_DB_10".Q;
   IF #_w1 THEN
       "OverspeedAlarm" := TRUE;
       "OverspeedNotify" := TRUE;
   END_IF;
   IF "AlarmReset" THEN "OvercurrentAlarm" := FALSE; END_IF;
   IF "AlarmSilence" OR "AlarmReset" THEN "OvercurrentNotify" := FALSE; END_IF;
END_REGION

REGION Network 5
   // High Oil Flow Alarm
   IF TRUE THEN
       #ti5 := "OilHighFlowDelay_Sp" * 1000;
       #tt5 := #ti5;
   END_IF;
   "IEC_Timer_0_DB_110".TON(IN := "OilFlow" > "OilHHflowSp", PT := #tt5);
   #_w1 := "IEC_Timer_0_DB_110".Q AND NOT #OS5;   // rising edge
   #OS5 := "IEC_Timer_0_DB_110".Q;
   IF #_w1 THEN
       "OilHighFlowAlarm" := TRUE;
       "OilHighFlowNotify" := TRUE;
   END_IF;
   IF "AlarmReset" THEN "OilHighFlowAlarm" := FALSE; END_IF;
   IF "AlarmSilence" OR "AlarmReset" THEN "OilHighFlowNotify" := FALSE; END_IF;
END_REGION

REGION Network 6
   // Brake Failure Alarm
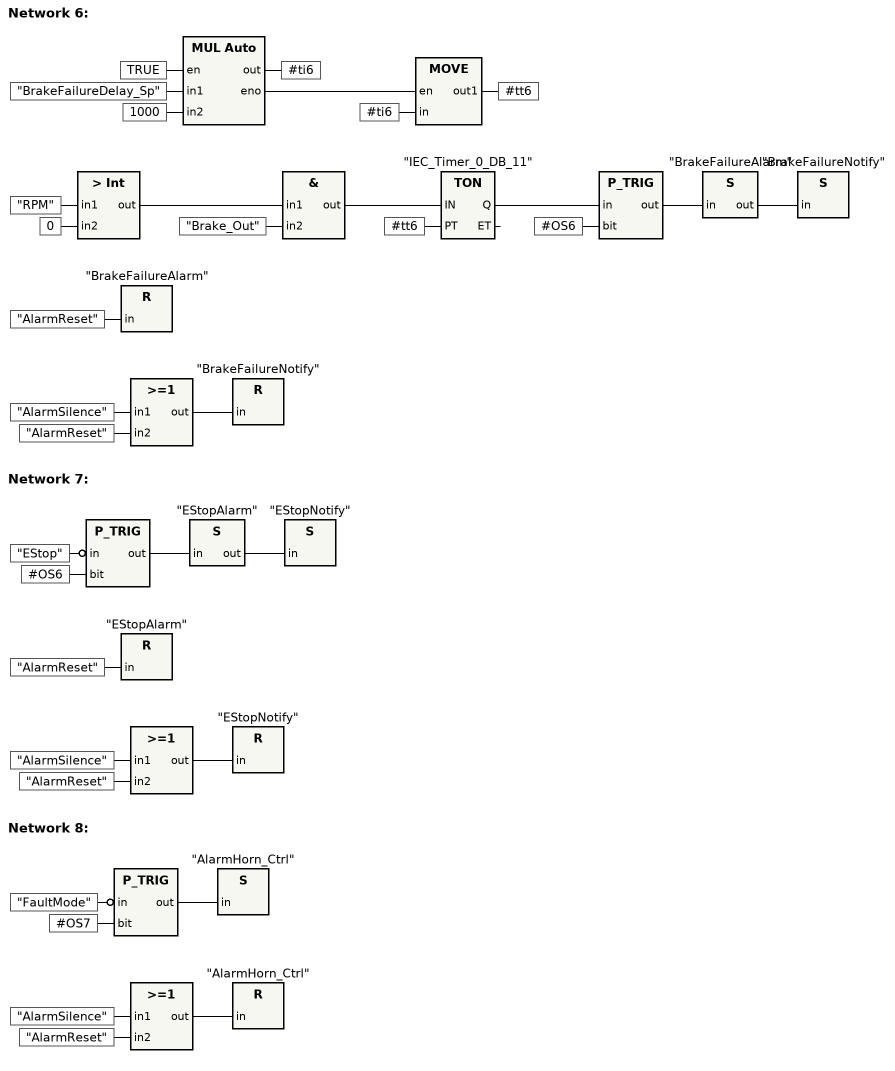
   IF TRUE THEN
       #ti6 := "BrakeFailureDelay_Sp" * 1000;
       #tt6 := #ti6;
   END_IF;
   "IEC_Timer_0_DB_11".TON(IN := ("RPM" > 0) AND "Brake_Out", PT := #tt6);
   #_w1 := "IEC_Timer_0_DB_11".Q AND NOT #OS6;   // rising edge
   #OS6 := "IEC_Timer_0_DB_11".Q;
   IF #_w1 THEN
       "BrakeFailureAlarm" := TRUE;
       "BrakeFailureNotify" := TRUE;
   END_IF;
   IF "AlarmReset" THEN "BrakeFailureAlarm" := FALSE; END_IF;
   IF "AlarmSilence" OR "AlarmReset" THEN "BrakeFailureNotify" := FALSE; END_IF;
END_REGION

REGION Network 7
   // EStop Alarm
   #_w1 := NOT "EStop" AND NOT #OS6;   // rising edge
   #OS6 := NOT "EStop";
   IF #_w1 THEN
       "EStopAlarm" := TRUE;
       "EStopNotify" := TRUE;
   END_IF;
   IF "AlarmReset" THEN "EStopAlarm" := FALSE; END_IF;
   IF "AlarmSilence" OR "AlarmReset" THEN "EStopNotify" := FALSE; END_IF;
END_REGION

REGION Network 8
   // Alarm Horn Control
   #_w1 := NOT "FaultMode" AND NOT #OS7;   // rising edge
   #OS7 := NOT "FaultMode";
   IF #_w1 THEN "AlarmHorn_Ctrl" := TRUE; END_IF;
   IF "AlarmSilence" OR "AlarmReset" THEN "AlarmHorn_Ctrl" := FALSE; END_IF;
END_REGION
END_FUNCTION_BLOCK

FUNCTION_BLOCK "ALARMS_SCL"   // FB12, SCL
{ S7_Optimized_Access := 'TRUE' }
VERSION : 0.1
   VAR_TEMP
      ti1 : Time;
      LOFAT : Bool;
      t1 : Time;
      ti2 : Time;
      ti3 : Time;
      ti4 : Time;
      ti5 : Time;
      ti6 : Time;
      ti7 : Time;
      t2 : Time;
      t3 : Time;
      t4 : Time;
      t5 : Time;
      t6 : Time;
      t7 : Time;
      OCAT : Bool;
      HOTAT : Bool;
      OSAT : Bool;
      HOFAT : Bool;
      BFAT : Bool;
   END_VAR
BEGIN
   //Oil Low Flow Alarm
   IF "OilPumpVFDen_Out" AND "OilFlow" < "OilLLflowSp" AND NOT "Brake_Out" AND NOT "OilLowFlowAlarm" AND NOT "AlarmReset" THEN
       "CONVERTTIME"(Int1 := "OilLowFlowDelay_Sp",
                     Time1 => #ti1);

       "IEC_Timer_0_DB_12".TON(IN := TRUE,
                               PT := #ti1,
                               Q => #LOFAT,
                               ET => #t1);
   END_IF;

   IF #LOFAT THEN
       "OilLowFlowAlarm" := 1;
       "OilLowFlowNotify" := 1;
   END_IF;

   IF "OilLowFlowAlarm" AND "AlarmReset" THEN
       "OilLowFlowAlarm" := 0;
       "OilLowFlowNotify" := 0;
   END_IF;

   IF "OilLowFlowNotify" AND "AlarmSilence" THEN
       "OilLowFlowNotify" := 0;
   END_IF;



   //Overcurrent Alarm
   IF "Current" > "OvercurrentSp" AND NOT "OvercurrentAlarm" AND NOT "AlarmReset" THEN
       "CONVERTTIME"(Int1:="OvercurrentDelay_Sp",
                     Time1=>#ti2);

       "IEC_Timer_0_DB_13".TON(IN:=TRUE,
                           PT:=#ti2,
                           Q=>#OCAT,
                           ET=>#t2);
   END_IF;

   IF #OCAT THEN
       "OvercurrentAlarm" := 1;
       "OvercurrentNotify" := 1;
   END_IF;

   IF "OvercurrentAlarm" AND "AlarmReset" THEN
       "OvercurrentAlarm" := 0;
       "OvercurrentNotify" := 0;
   END_IF;

   IF "OvercurrentNotify" AND "AlarmSilence" THEN
       "OvercurrentNotify" := 0;
   END_IF;




   //High Oil Temp Alarm
   IF "OilTemp" > "HighOilTempSp" AND NOT "HighOilTempAlarm" AND NOT "AlarmReset" THEN
       "CONVERTTIME"(Int1 := "HighOilTempDelay_Sp",
                     Time1 => #ti3);

   "IEC_Timer_0_DB_14".TON(IN:=TRUE,
                           PT:=#ti3,
                           Q=>#HOTAT,
                           ET=>#t3);
   END_IF;

   IF #HOTAT THEN
       "HighOilTempAlarm" := 1;
       "HighOilTempNotify" := 1;
   END_IF;

   IF "HighOilTempAlarm" AND "AlarmReset" THEN
       "HighOilTempAlarm" := 0;
       "HighOilTempNotify" := 0;
   END_IF;

   IF "HighOilTempNotify" AND "AlarmSilence" THEN
       "HighOilTempNotify" := 0;
   END_IF;



   //Overspeed Alarm
   IF "RPM" > "OverspeedSp" AND NOT "OverspeedAlarm" AND NOT "AlarmReset" THEN
   "CONVERTTIME"(Int1:="OverspeedDelay_Sp",
                 Time1=>#ti4);
   "IEC_Timer_0_DB_15".TON(IN:=TRUE,
                           PT:=#ti4,
                           Q=>#OSAT,
                           ET=>#t4);
   END_IF;

   IF #OSAT THEN
       "OverspeedAlarm" := 1;
       "OverspeedNotify" := 1;
   END_IF;

   IF "OverspeedAlarm" AND "AlarmReset" THEN
       "OverspeedAlarm" := 0;
       "OverspeedNotify" := 0;
   END_IF;

   IF "OverspeedNotify" AND "AlarmSilence" THEN
       "OverspeedNotify" := 0;
   END_IF;



   //High Oil Flow Alarm
   IF "OilFlow" > "OilHHflowSp" AND NOT "OilHighFlowAlarm" AND NOT "AlarmReset" THEN
   "CONVERTTIME"(Int1:="OilHighFlowDelay_Sp",
                 Time1=>#ti5);
   "IEC_Timer_0_DB_16".TON(IN:=TRUE,
                           PT:=#ti5,
                           Q=>#HOFAT,
                           ET=>#t5);

   END_IF;

   IF #HOFAT THEN
       "OilHighFlowAlarm" := 1;
       "OilHighFlowNotify" := 1;
   END_IF;

   IF "OilHighFlowAlarm" AND "AlarmReset" THEN
       "OilHighFlowAlarm" := 0;
       "OilHighFlowNotify" := 0;
   END_IF;

   IF "OilHighFlowNotify" AND "AlarmSilence" THEN
       "OilHighFlowNotify" := 0;
   END_IF;



   //Brake Failure Alarm
   IF "Brake_Out" AND "RPM" > 0 AND NOT "BrakeFailureAlarm" AND NOT "AlarmReset" THEN
   "CONVERTTIME"(Int1:="BrakeFailureDelay_Sp",
                 Time1=>#ti6);
   "IEC_Timer_0_DB_17".TON(IN:=TRUE,
                           PT:=#ti6,
                           Q=>#BFAT,
                           ET=>#t6);
   END_IF;

   IF #BFAT THEN
       "BrakeFailureAlarm" := 1;
       "BrakeFailureNotify" := 1;
   END_IF;

   IF "BrakeFailureAlarm" AND "AlarmReset" THEN
       "BrakeFailureAlarm" := 0;
       "BrakeFailureNotify" := 0;
   END_IF;

   IF "BrakeFailureNotify" AND "AlarmSilence" THEN
       "BrakeFailureNotify" := 0;
   END_IF;

